screen "40_SimValues_5" 800x480, template "31_SimValues_1"
   GraphicView "gfxDarkBackground" at 0,0 size 800x480; Picture "PopUpBackground"
      Visibility <- "PopUpBackground"
   TextField "txtParameter1_2" at 246,136 size 42x25; Text 'Step 2 / Parameter 1'
   TextField "txtParameter1_3" at 316,136 size 102x25; Text 'Step 3 / Parameter 1'
   TextField "txtParameter1_4" at 386,136 size 102x25; Text 'Step 4 / Parameter 1'
   TextField "txtParameter1_5" at 456,136 size 102x25; Text 'Step 5 / Parameter 1'
   TextField "txtParameter1_6" at 526,136 size 102x25; Text 'Step 6 / Parameter 1'
   TextField "txtParameter1_8" at 596,136 size 102x25; Text 'Step 7 / Parameter 1'
   TextField "txtParameter1_9" at 666,136 size 102x25; Text 'Step 8 / Parameter 1'
   TextField "txtParameter1_10" at 176,136 size 45x25; Text 'Step 1 / Parameter 1'
   TextField "txtParameter1_11" at 736,136 size 46x25; Text 'Step 9 / Parameter 1'
   TextField "txtParameter1_1" at 104,136 size 45x25; Text 'Branch / Parameter 1'
   TextField "txtParameter1_7" at 32,136 size 45x25; Text 'Car / Parameter 1'
   GraphicView "Graphic view_1" at 33,184 size 40x40; Picture "Car_Red"
   GraphicView "Graphic view_3" at 33,249 size 40x40; Picture "Car_Green"
   GraphicView "Graphic view_4" at 33,308 size 40x40; Picture "Car_Blue_1"
   TextField "Text field_3" at 121,191 size 15x23; Text '1'
      Visibility <- "InScreenTabState"
   TextField "Text field_1" at 121,256 size 15x23; Text '2'
      Visibility <- "InScreenTabState"
   TextField "Text field_2" at 121,321 size 15x23; Text '2'
      Visibility <- "InScreenTabState"
   Button "Button_1" at 176,186 size 38x32; TextOff 'Text'
      on Click: SetTag("DB_HMI_ARG1_Seq1_DelaySelect_Red{2}(4)", 1)
   Button "Button_2" at 245,186 size 38x32; TextOff 'Text'
      on Click: SetTag("DB_HMI_ARG1_Seq1_DelaySelect_Red{3}(4)", 1)
   Button "Button_3" at 315,186 size 38x32; TextOff 'Text'
      on Click: SetTag("DB_HMI_ARG1_Seq1_DelaySelect_Red{4}(4)", 1)
   Button "Button_4" at 385,186 size 38x32; TextOff 'Text'
      on Click: SetTag("DB_HMI_ARG1_Seq1_DelaySelect_Red{5}(4)", 1)
   Button "Button_5" at 455,186 size 38x32; TextOff 'Text'
      on Click: SetTag("DB_HMI_ARG1_Seq1_DelaySelect_Red{6}(4)", 1)
   Button "Button_6" at 525,186 size 38x32; TextOff 'Text'
      on Click: SetTag("DB_HMI_ARG1_Seq1_DelaySelect_Red{7}(4)", 1)
   Button "Button_8" at 595,186 size 38x32; TextOff 'Text'
      on Click: SetTag("DB_HMI_ARG1_Seq1_DelaySelect_Red{8}(4)", 1)
   Button "Button_9" at 665,186 size 38x32; TextOff 'Text'
      on Click: SetTag("DB_HMI_ARG1_Seq1_DelaySelect_Red{9}(4)", 1)
   Button "Button_10" at 735,186 size 38x32; TextOff 'Text'
      on Click: SetTag("DB_HMI_ARG1_Seq1_DelaySelect_Red{10}(4)", 1)
   Button "Button_17" at 176,250 size 38x32; TextOff 'Text'
      on Click: SetTag("DB_HMI_ARG1_Seq1_DelaySelect_Green{2}(4)", 1)
   Button "Button_7" at 246,250 size 38x32; TextOff 'Text'
      on Click: SetTag("DB_HMI_ARG1_Seq1_DelaySelect_Green{3}(4)", 1)
   Button "Button_11" at 316,250 size 38x32; TextOff 'Text'
      on Click: SetTag("DB_HMI_ARG1_Seq1_DelaySelect_Green{4}(4)", 1)
   Button "Button_12" at 386,250 size 38x32; TextOff 'Text'
      on Click: SetTag("DB_HMI_ARG1_Seq1_DelaySelect_Green{5}(4)", 1)
   Button "Button_13" at 456,250 size 38x32; TextOff 'Text'
      on Click: SetTag("DB_HMI_ARG1_Seq1_DelaySelect_Green{6}(4)", 1)
   Button "Button_14" at 526,250 size 38x32; TextOff 'Text'
      on Click: SetTag("DB_HMI_ARG1_Seq1_DelaySelect_Green{7}(4)", 1)
   Button "Button_15" at 596,250 size 38x32; TextOff 'Text'
      on Click: SetTag("DB_HMI_ARG1_Seq1_DelaySelect_Green{8}(4)", 1)
   Button "Button_16" at 666,250 size 38x32; TextOff 'Text'
      on Click: SetTag("DB_HMI_ARG1_Seq1_DelaySelect_Green{9}(4)", 1)
   Button "Button_18" at 736,250 size 38x32; TextOff 'Text'
      on Click: SetTag("DB_HMI_ARG1_Seq1_DelaySelect_Green{10}(4)", 1)
   Button "Button_26" at 176,314 size 38x32; TextOff 'Text'
      on Click: SetTag("DB_HMI_ARG1_Seq1_DelaySelect_Blue{2}(4)", 1)
   Button "Button_19" at 246,314 size 38x32; TextOff 'Text'
      on Click: SetTag("DB_HMI_ARG1_Seq1_DelaySelect_Blue{3}(4)", 1)
   Button "Button_20" at 316,314 size 38x32; TextOff 'Text'
      on Click: SetTag("DB_HMI_ARG1_Seq1_DelaySelect_Blue{4}(4)", 1)
   Button "Button_21" at 386,314 size 38x32; TextOff 'Text'
      on Click: SetTag("DB_HMI_ARG1_Seq1_DelaySelect_Blue{5}(4)", 1)
   Button "Button_22" at 456,314 size 38x32; TextOff 'Text'
      on Click: SetTag("DB_HMI_ARG1_Seq1_DelaySelect_Blue{6}(4)", 1)
   Button "Button_23" at 526,314 size 38x32; TextOff 'Text'
      on Click: SetTag("DB_HMI_ARG1_Seq1_DelaySelect_Blue{7}(4)", 1)
   Button "Button_24" at 596,314 size 38x32; TextOff 'Text'
      on Click: SetTag("DB_HMI_ARG1_Seq1_DelaySelect_Blue{8}(4)", 1)
   Button "Button_25" at 666,314 size 38x32; TextOff 'Text'
      on Click: SetTag("DB_HMI_ARG1_Seq1_DelaySelect_Blue{9}(4)", 1)
   Button "Button_27" at 736,314 size 38x32; TextOff 'Text'
      on Click: SetTag("DB_HMI_ARG1_Seq1_DelaySelect_Blue{10}(4)", 1)
   Button "Button_28" at 176,186 size 38x32; TextOff 'Text'
      on Click: SetTag("DB_HMI_ARG1_Seq1_DelaySelect_Red{2}(4)", 0)
      Visibility <- "DB_HMI_ARG1_Seq1_DelaySelect_Red{2}(4)"
   Button "Button_29" at 245,186 size 38x32; TextOff 'Text'
      on Click: SetTag("DB_HMI_ARG1_Seq1_DelaySelect_Red{3}(4)", 0)
      Visibility <- "DB_HMI_ARG1_Seq1_DelaySelect_Red{3}(4)"
   Button "Button_30" at 315,186 size 38x32; TextOff 'Text'
      on Click: SetTag("DB_HMI_ARG1_Seq1_DelaySelect_Red{4}(4)", 0)
      Visibility <- "DB_HMI_ARG1_Seq1_DelaySelect_Red{4}(4)"
   Button "Button_31" at 385,186 size 38x32; TextOff 'Text'
      on Click: SetTag("DB_HMI_ARG1_Seq1_DelaySelect_Red{5}(4)", 0)
      Visibility <- "DB_HMI_ARG1_Seq1_DelaySelect_Red{5}(4)"
   Button "Button_32" at 455,186 size 38x32; TextOff 'Text'
      on Click: SetTag("DB_HMI_ARG1_Seq1_DelaySelect_Red{6}(4)", 0)
      Visibility <- "DB_HMI_ARG1_Seq1_DelaySelect_Red{6}(4)"
   Button "Button_33" at 525,186 size 38x32; TextOff 'Text'
      on Click: SetTag("DB_HMI_ARG1_Seq1_DelaySelect_Red{7}(4)", 0)
      Visibility <- "DB_HMI_ARG1_Seq1_DelaySelect_Red{7}(4)"
   Button "Button_34" at 595,186 size 38x32; TextOff 'Text'
      on Click: SetTag("DB_HMI_ARG1_Seq1_DelaySelect_Red{8}(4)", 0)
      Visibility <- "DB_HMI_ARG1_Seq1_DelaySelect_Red{8}(4)"
   Button "Button_35" at 665,186 size 38x32; TextOff 'Text'
      on Click: SetTag("DB_HMI_ARG1_Seq1_DelaySelect_Red{9}(4)", 0)
      Visibility <- "DB_HMI_ARG1_Seq1_DelaySelect_Red{9}(4)"
   Button "Button_36" at 735,186 size 38x32; TextOff 'Text'
      on Click: SetTag("DB_HMI_ARG1_Seq1_DelaySelect_Red{10}(4)", 0)
      Visibility <- "DB_HMI_ARG1_Seq1_DelaySelect_Red{10}(4)"
   Button "Button_37" at 176,250 size 38x32; TextOff 'Text'
      on Click: SetTag("DB_HMI_ARG1_Seq1_DelaySelect_Green{2}(4)", 0)
      Visibility <- "DB_HMI_ARG1_Seq1_DelaySelect_Green{2}(4)"
   Button "Button_38" at 246,250 size 38x32; TextOff 'Text'
      on Click: SetTag("DB_HMI_ARG1_Seq1_DelaySelect_Green{3}(4)", 0)
      Visibility <- "DB_HMI_ARG1_Seq1_DelaySelect_Green{3}(4)"
   Button "Button_39" at 316,250 size 38x32; TextOff 'Text'
      on Click: SetTag("DB_HMI_ARG1_Seq1_DelaySelect_Green{4}(4)", 0)
      Visibility <- "DB_HMI_ARG1_Seq1_DelaySelect_Green{4}(4)"
   Button "Button_40" at 386,250 size 38x32; TextOff 'Text'
      on Click: SetTag("DB_HMI_ARG1_Seq1_DelaySelect_Green{5}(4)", 0)
      Visibility <- "DB_HMI_ARG1_Seq1_DelaySelect_Green{5}(4)"
   Button "Button_41" at 456,250 size 38x32; TextOff 'Text'
      on Click: SetTag("DB_HMI_ARG1_Seq1_DelaySelect_Green{6}(4)", 0)
      Visibility <- "DB_HMI_ARG1_Seq1_DelaySelect_Green{6}(4)"
   Button "Button_42" at 526,250 size 38x32; TextOff 'Text'
      on Click: SetTag("DB_HMI_ARG1_Seq1_DelaySelect_Green{7}(4)", 0)
      Visibility <- "DB_HMI_ARG1_Seq1_DelaySelect_Green{7}(4)"
   Button "Button_43" at 596,250 size 38x32; TextOff 'Text'
      on Click: SetTag("DB_HMI_ARG1_Seq1_DelaySelect_Green{8}(4)", 0)
      Visibility <- "DB_HMI_ARG1_Seq1_DelaySelect_Green{8}(4)"
   Button "Button_44" at 666,250 size 38x32; TextOff 'Text'
      on Click: SetTag("DB_HMI_ARG1_Seq1_DelaySelect_Green{9}(4)", 0)
      Visibility <- "DB_HMI_ARG1_Seq1_DelaySelect_Green{9}(4)"
   Button "Button_45" at 736,250 size 38x32; TextOff 'Text'
      on Click: SetTag("DB_HMI_ARG1_Seq1_DelaySelect_Green{10}(4)", 0)
      Visibility <- "DB_HMI_ARG1_Seq1_DelaySelect_Green{10}(4)"
   Button "Button_46" at 176,314 size 38x32; TextOff 'Text'
      on Click: SetTag("DB_HMI_ARG1_Seq1_DelaySelect_Blue{2}(4)", 0)
      Visibility <- "DB_HMI_ARG1_Seq1_DelaySelect_Blue{2}(4)"
   Button "Button_47" at 246,314 size 38x32; TextOff 'Text'
      on Click: SetTag("DB_HMI_ARG1_Seq1_DelaySelect_Blue{3}(4)", 0)
      Visibility <- "DB_HMI_ARG1_Seq1_DelaySelect_Blue{3}(4)"
   Button "Button_48" at 316,314 size 38x32; TextOff 'Text'
      on Click: SetTag("DB_HMI_ARG1_Seq1_DelaySelect_Blue{4}(4)", 0)
      Visibility <- "DB_HMI_ARG1_Seq1_DelaySelect_Blue{4}(4)"
   Button "Button_49" at 386,314 size 38x32; TextOff 'Text'
      on Click: SetTag("DB_HMI_ARG1_Seq1_DelaySelect_Blue{5}(4)", 0)
      Visibility <- "DB_HMI_ARG1_Seq1_DelaySelect_Blue{5}(4)"
   Button "Button_50" at 456,314 size 38x32; TextOff 'Text'
      on Click: SetTag("DB_HMI_ARG1_Seq1_DelaySelect_Blue{6}(4)", 0)
      Visibility <- "DB_HMI_ARG1_Seq1_DelaySelect_Blue{6}(4)"
   Button "Button_51" at 526,314 size 38x32; TextOff 'Text'
      on Click: SetTag("DB_HMI_ARG1_Seq1_DelaySelect_Blue{7}(4)", 0)
      Visibility <- "DB_HMI_ARG1_Seq1_DelaySelect_Blue{7}(4)"
   Button "Button_52" at 596,314 size 38x32; TextOff 'Text'
      on Click: SetTag("DB_HMI_ARG1_Seq1_DelaySelect_Blue{8}(4)", 0)
      Visibility <- "DB_HMI_ARG1_Seq1_DelaySelect_Blue{8}(4)"
   Button "Button_53" at 666,314 size 38x32; TextOff 'Text'
      on Click: SetTag("DB_HMI_ARG1_Seq1_DelaySelect_Blue{9}(4)", 0)
      Visibility <- "DB_HMI_ARG1_Seq1_DelaySelect_Blue{9}(4)"
   Button "Button_54" at 736,314 size 38x32; TextOff 'Text'
      on Click: SetTag("DB_HMI_ARG1_Seq1_DelaySelect_Blue{10}(4)", 0)
      Visibility <- "DB_HMI_ARG1_Seq1_DelaySelect_Blue{10}(4)"
   Button "Button_55" at 619,378 size 165x40; TextOff 'Reset / Alle Quittieren'; PictureOff "More_Icon"
      on ReleaseLeft: ResetBit("Ext_AckSafety_DB_ack")
      on PressLeft: SetBit("Ext_AckSafety_DB_ack")
      on Release: SetTag("DB_HMI_ARG1_Seq1_Cmd_DelayReset(4)", 0)
      on Press: SetTag("DB_HMI_ARG1_Seq1_Cmd_DelayReset(4)", 1)
      ObjectEnable <- "DB_HMI_ARG1_Seq1_Cmd_DelayReset"

Template "01_Navigation" 800x480
   Gauge "gaugeDiagStateUpdate" at 566,2 size 50x50; CaptionText 'SIMATIC'
      ProcessValue <- "@DiagnosticsIndicatorTag"
   TextField "txtTitleBar" at 16,8 size 495x32; Text 'Step Time Analysis / Applikation'
   Button "btnSubNavActive1" at 0,432 size 133x48; TextOff 'Overview / Übersicht'
      Visibility <- "SubNavigationState"
   Button "btnSubNavActive2" at 133,432 size 133x48; TextOff 'Station 1 / Modul 1'
      Visibility <- "SubNavigationState"
   Button "btnSubNavActive3" at 266,432 size 133x48; TextOff 'Station 2 / Modul 2'
      Visibility <- "SubNavigationState"
   Button "btnSubNavActive4" at 399,432 size 133x48; TextOff 'Station 3 / Modul 3'
      Visibility <- "SubNavigationState"
   Button "btnSubNavActive5" at 532,432 size 133x48; TextOff 'Station 4 / Modul 4'
      Visibility <- "SubNavigationState"
   Button "btnSubNavActive5_1" at 665,432 size 133x48; TextOff 'Station 5 / Modul 4'
      Visibility <- "SubNavigationState"
   Rectangle "rectIndicatorActive1" at 0,475 size 133x5
      Visibility <- "SubNavigationState"
   Rectangle "rectIndicatorActive2" at 133,475 size 133x5
      Visibility <- "SubNavigationState"
   Rectangle "rectIndicatorActive3" at 266,475 size 133x5
      Visibility <- "SubNavigationState"
   Rectangle "rectIndicatorActive4" at 399,475 size 133x5
      Visibility <- "SubNavigationState"
   Rectangle "rectIndicatorActive5" at 532,475 size 133x5
      Visibility <- "SubNavigationState"
   Rectangle "rectIndicatorActive5_1" at 665,475 size 133x5
      Visibility <- "SubNavigationState"
   GraphicView "gfxPrevScreenIcon" at 704,444 size 24x24; Picture "PrevScreen_Icon"
   Button "btnSubNav1" at 0,432 size 133x48; TextOff 'Overview / Übersicht'
      on Click: SetTag("SubNavigationState", 1); ActivateScreen("10_Startscreen", 0)
   Button "btnSubNav2" at 133,432 size 133x48; TextOff 'Station 1 / Modul 1'
      on Click: SetTag("SubNavigationState", 2); ActivateScreen("21_Station_1", 0)
   Button "btnSubNav3" at 266,432 size 133x48; TextOff 'Station 2 / Modul 2'
      on Click: SetTag("SubNavigationState", 3); ActivateScreen("22_Station_2", 0)
   Button "btnSubNav4" at 399,432 size 133x48; TextOff 'Station 3 / Modul 3'
      on Click: SetTag("SubNavigationState", 4); ActivateScreen("23_Station_3", 0)
   Button "btnSubNav5" at 532,432 size 133x48; TextOff 'Station 4 / Modul 4'
      on Click: SetTag("SubNavigationState", 5); ActivateScreen("24_Station_4", 0)
   Button "btnSubNav6" at 665,432 size 135x48; TextOff 'Station 5 / Modul 4'
      on Click: SetTag("SubNavigationState", 6); ActivateScreen("25_Station_5", 0)
   Button "btnStartscreen" at 0,0 size 250x45; TextOff 'Text'
      on Click: ActivateScreen("10_Startscreen", 0)

Template "21_Station_1" 800x480
   Gauge "gaugeDiagStateUpdate" at 566,2 size 50x50; CaptionText 'SIMATIC'
      ProcessValue <- "@DiagnosticsIndicatorTag"
   TextField "txtTitleBar" at 16,8 size 495x32; Text 'Step Time Analysis / Applikation'
   Button "btnSubNavActive1" at 0,432 size 133x48; TextOff 'Overview / Übersicht'
      Visibility <- "SubNavigationState"
   Button "btnSubNavActive2" at 133,432 size 133x48; TextOff 'Station 1 / Modul 1'
      Visibility <- "SubNavigationState"
   Button "btnSubNavActive3" at 266,432 size 133x48; TextOff 'Station 2 / Modul 2'
      Visibility <- "SubNavigationState"
   Button "btnSubNavActive4" at 399,432 size 133x48; TextOff 'Station 3 / Modul 3'
      Visibility <- "SubNavigationState"
   Button "btnSubNavActive5" at 532,432 size 133x48; TextOff 'Station 4 / Modul 4'
      Visibility <- "SubNavigationState"
   Button "btnSubNavActive5_1" at 665,432 size 133x48; TextOff 'Station 5 / Modul 4'
      Visibility <- "SubNavigationState"
   Rectangle "rectIndicatorActive1" at 0,475 size 133x5
      Visibility <- "SubNavigationState"
   Rectangle "rectIndicatorActive2" at 133,475 size 133x5
      Visibility <- "SubNavigationState"
   Rectangle "rectIndicatorActive3" at 266,475 size 133x5
      Visibility <- "SubNavigationState"
   Rectangle "rectIndicatorActive4" at 399,475 size 133x5
      Visibility <- "SubNavigationState"
   Rectangle "rectIndicatorActive5" at 532,475 size 133x5
      Visibility <- "SubNavigationState"
   Rectangle "rectIndicatorActive5_1" at 665,475 size 133x5
      Visibility <- "SubNavigationState"
   GraphicView "gfxPrevScreenIcon" at 704,444 size 24x24; Picture "PrevScreen_Icon"
   Button "btnSubNav1" at 0,432 size 133x48; TextOff 'Overview / Übersicht'
      on Click: SetTag("SubNavigationState", 1); ActivateScreen("10_Startscreen", 0)
   Button "btnSubNav2" at 133,432 size 133x48; TextOff 'Station 1 / Modul 1'
      on Click: SetTag("SubNavigationState", 2); ActivateScreen("21_Station_1", 0)
   Button "btnSubNav3" at 266,432 size 133x48; TextOff 'Station 2 / Modul 2'
      on Click: SetTag("SubNavigationState", 3); ActivateScreen("22_Station_2", 0)
   Button "btnSubNav4" at 399,432 size 133x48; TextOff 'Station 3 / Modul 3'
      on Click: SetTag("SubNavigationState", 4); ActivateScreen("23_Station_3", 0)
   Button "btnSubNav5" at 532,432 size 133x48; TextOff 'Station 4 / Modul 4'
      on Click: SetTag("SubNavigationState", 5); ActivateScreen("24_Station_4", 0)
   Button "btnSubNav6" at 665,432 size 135x48; TextOff 'Station 5 / Modul 4'
      on Click: SetTag("SubNavigationState", 6); ActivateScreen("25_Station_5", 0)
   Button "btnStartscreen" at 0,0 size 250x45; TextOff 'Text'
      on Click: ActivateScreen("10_Startscreen", 0)
   Rectangle "rectState" at 0,48 size 56x38
      Appearance <- "CurrentMachineState"
   Button "btnState" at 201,53 size 34x31; TextOff '...'; PictureOff "More_Icon"
      on Click: ActivateScreen("31_Mode_Station_1", 0)
   TextField "Auto" at 67,63 size 34x19; Text 'Auto'
      Visibility <- "DB_HMI_ARG1_Seq1_Status_Auto"
   TextField "Manual" at 69,63 size 31x19; Text 'Man'
      Visibility <- "DB_HMI_ARG1_Seq1_Status_Man"
   TextField "txtStateHeadline" at 65,48 size 123x23; Text 'Mode / Status'

Template "31_SimValues_1" 800x480
   Gauge "gaugeDiagStateUpdate" at 566,2 size 50x50; CaptionText 'SIMATIC'
      ProcessValue <- "@DiagnosticsIndicatorTag"
   TextField "txtTitleBar" at 16,8 size 495x32; Text 'Step Time Analysis / Applikation'
   GraphicView "gfxPrevScreenIcon" at 704,444 size 24x24; Picture "PrevScreen_Icon"
   GraphicView "gfxPrevScreenIcon_1" at 705,444 size 24x24; Picture "PrevScreen_Icon"
   Button "btnPreviousScreen" at 688,432 size 56x48; TextOff 'Text'
      on Click: function_efd93a16()
   Button "btnStartscreen" at 0,0 size 250x45; TextOff 'Text'
      on Click: ActivateScreen("10_Startscreen", 0)

VB script "movingCar"
   'Tip:
   ' 1. Use the <CTRL+SPACE> or <CTRL+I> shortcut to open a list of all objects and functions
   ' 2. Write the code using the HMI Runtime object.
   '  Example: HmiRuntime.Screens("Screen_1").
   ' 3. Use the <CTRL+J> shortcut to create an object reference.
   'Write the code as of this position:
   
   'car movement
   
   'Please replace all sequences which are enclosed with '_' by your own code.
   
   If SmartTags("DB_HMI_ARG1_Seq1_S1") = True Then
   	SmartTags("StepNumber")= 0                                            
   End If 
   
   If SmartTags("DB_HMI_ARG1_Seq1_S2") = True Or SmartTags("DB_HMI_ARG1_Seq1_S11") = True Then
   	SmartTags("StepNumber")= 1                                            
   End If                                                                    
   If SmartTags("DB_HMI_ARG1_Seq1_S3") = True Or SmartTags("DB_HMI_ARG1_Seq1_S12") = True Then
   	SmartTags("StepNumber")= 2                                            
   End If                                                                    
   If SmartTags("DB_HMI_ARG1_Seq1_S4") = True Or SmartTags("DB_HMI_ARG1_Seq1_S13") = True Then
   	SmartTags("StepNumber")= 3                                            
   End If                                                                    
   If SmartTags("DB_HMI_ARG1_Seq1_S5") = True Or SmartTags("DB_HMI_ARG1_Seq1_S14") = True Then
   	SmartTags("StepNumber")= 4                                            
   End If                                                                    
   If SmartTags("DB_HMI_ARG1_Seq1_S6") = True Or SmartTags("DB_HMI_ARG1_Seq1_S15") = True Then
   	SmartTags("StepNumber")= 5                                            
   End If                                                                    
   If SmartTags("DB_HMI_ARG1_Seq1_S7") = True Or SmartTags("DB_HMI_ARG1_Seq1_S16") = True Then
   	SmartTags("StepNumber")= 6                                            
   End If                                                                    
   If SmartTags("DB_HMI_ARG1_Seq1_S8") = True Or SmartTags("DB_HMI_ARG1_Seq1_S17") = True Then
   	SmartTags("StepNumber")= 7                                            
   End If                                                                    
   If SmartTags("DB_HMI_ARG1_Seq1_S9") = True Or SmartTags("DB_HMI_ARG1_Seq1_S18") = True Then
   	SmartTags("StepNumber")= 8                                             
   End If                                                                     
   If SmartTags("DB_HMI_ARG1_Seq1_S10") = True Or SmartTags("DB_HMI_ARG1_Seq1_S19") = True Then
   	SmartTags("StepNumber")= 9                 
   End If                                         

VB script "VBFunction_1"
   'Tip:
   ' 1. Use the <CTRL+SPACE> or <CTRL+I> shortcut to open a list of all objects and functions
   ' 2. Write the code using the HMI Runtime object.
   '  Example: HmiRuntime.Screens("Screen_1").
   ' 3. Use the <CTRL+J> shortcut to create an object reference.
   'Write the code as of this position:
   
   
   'Please replace all sequences which are enclosed with '_' by your own code.
   If SmartTags("DB_HMI_ARG1_Seq1_Status_Idle")=True Then
   	SmartTags("status")=0
   ElseIf SmartTags("DB_HMI_ARG1_Seq1_Status_Busy")= True Then
   	SmartTags("status")=1
   Else
   	SmartTags("status")=2
   End If

scheduled task "UserName"
   on Action: function_f41c6f6c("CurrentUserName")
*)